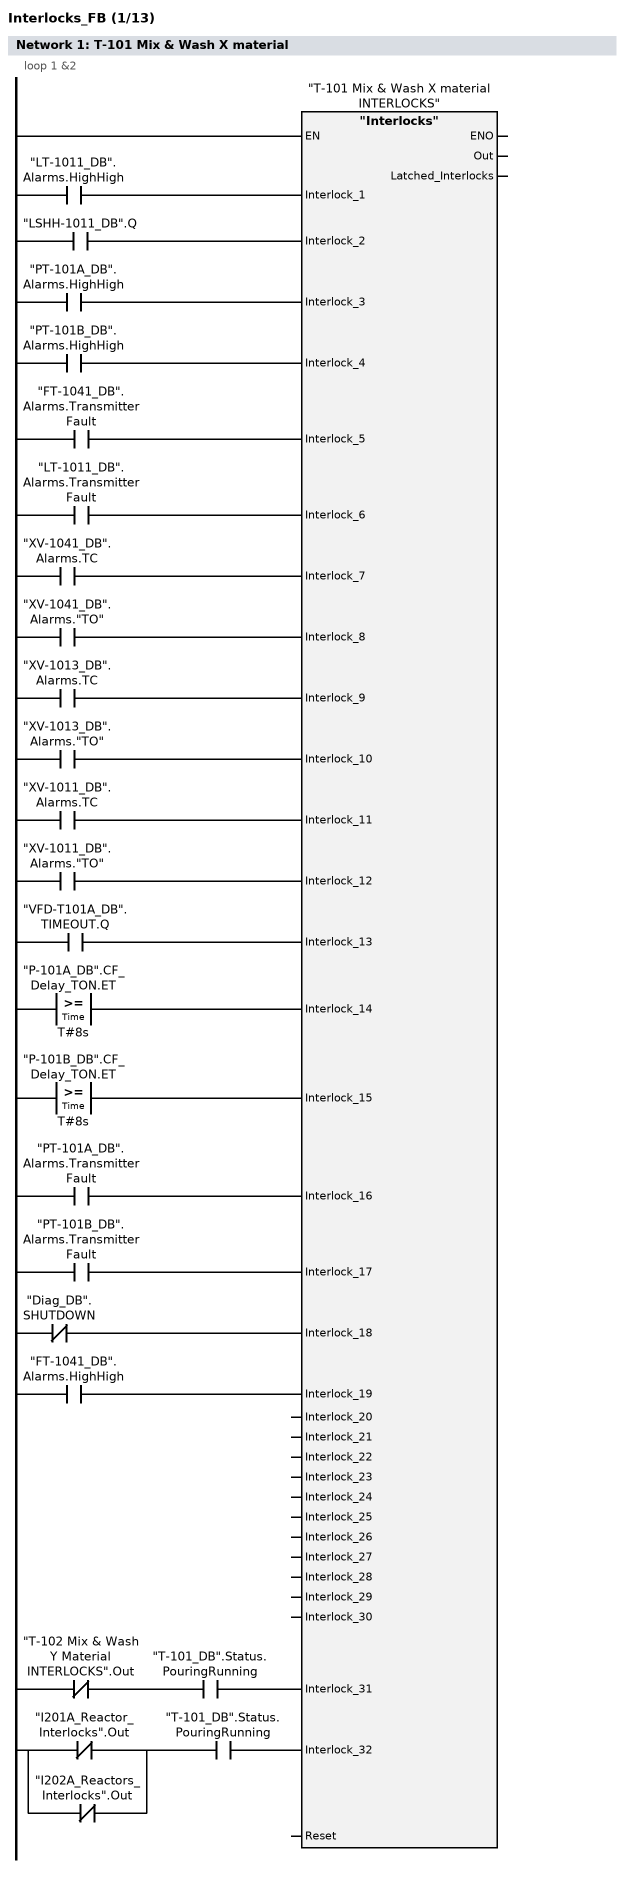
   RUNG wire#powerrail
      "T-101 Mix & Wash X material INTERLOCKS"(Interlock_1 := wire#w1, Interlock_2 := wire#w2, Interlock_3 := wire#w3, Interlock_4 := wire#w4, Interlock_5 := wire#w5, Interlock_6 := wire#w6, Interlock_7 := wire#w7, Interlock_8 := wire#w8, Interlock_9 := wire#w9, Interlock_10 := wire#w10, Interlock_11 := wire#w11, Interlock_12 := wire#w12, Interlock_13 := wire#w13, Interlock_14 := wire#w14, Interlock_15 := wire#w15, Interlock_16 := wire#w16, Interlock_17 := wire#w17, Interlock_18 := wire#w18, Interlock_19 := wire#w19, Interlock_31 := wire#w20, Interlock_32 := wire#w22, Interlock_20 :=, Interlock_21 :=, Interlock_22 :=, Interlock_23 :=, Interlock_24 :=, Interlock_25 :=, Interlock_26 :=, Interlock_27 :=, Interlock_28 :=, Interlock_29 :=, Interlock_30 :=, Reset :=, Out =>, Latched_Interlocks =>)
   END_RUNG
   RUNG wire#powerrail
      Contact( "LT-1011_DB".Alarms.HighHigh )
   END_RUNG wire#w1
   RUNG wire#powerrail
      Contact( "LSHH-1011_DB".Q )
   END_RUNG wire#w2
   RUNG wire#powerrail
      Contact( "PT-101A_DB".Alarms.HighHigh )
   END_RUNG wire#w3
   RUNG wire#powerrail
      Contact( "PT-101B_DB".Alarms.HighHigh )
   END_RUNG wire#w4
   RUNG wire#powerrail
      Contact( "FT-1041_DB".Alarms.TransmitterFault )
   END_RUNG wire#w5
   RUNG wire#powerrail
      Contact( "LT-1011_DB".Alarms.TransmitterFault )
   END_RUNG wire#w6
   RUNG wire#powerrail
      Contact( "XV-1041_DB".Alarms.TC )
   END_RUNG wire#w7
   RUNG wire#powerrail
      Contact( "XV-1041_DB".Alarms."TO" )
   END_RUNG wire#w8
   RUNG wire#powerrail
      Contact( "XV-1013_DB".Alarms.TC )
   END_RUNG wire#w9
   RUNG wire#powerrail
      Contact( "XV-1013_DB".Alarms."TO" )
   END_RUNG wire#w10
   RUNG wire#powerrail
      Contact( "XV-1011_DB".Alarms.TC )
   END_RUNG wire#w11
   RUNG wire#powerrail
      Contact( "XV-1011_DB".Alarms."TO" )
   END_RUNG wire#w12
   RUNG wire#powerrail
      Contact( "VFD-T101A_DB".TIMEOUT.Q )
   END_RUNG wire#w13
   RUNG wire#powerrail
      { S7_Templates := "SrcType := Time" } GE_Contact(in1 := "P-101A_DB".CF_Delay_TON.ET, in2 := T#8s)
   END_RUNG wire#w14
   RUNG wire#powerrail
      { S7_Templates := "SrcType := Time" } GE_Contact(in1 := "P-101B_DB".CF_Delay_TON.ET, in2 := T#8s)
   END_RUNG wire#w15
   RUNG wire#powerrail
      Contact( "PT-101A_DB".Alarms.TransmitterFault )
   END_RUNG wire#w16
   RUNG wire#powerrail
      Contact( "PT-101B_DB".Alarms.TransmitterFault )
   END_RUNG wire#w17
   RUNG wire#powerrail
      I_Contact( "Diag_DB".SHUTDOWN )
   END_RUNG wire#w18
   RUNG wire#powerrail
      Contact( "FT-1041_DB".Alarms.HighHigh )
   END_RUNG wire#w19
   RUNG wire#powerrail
      I_Contact( "T-102 Mix & Wash Y Material  INTERLOCKS".Out )
      Contact( "T-101_DB".Status.PouringRunning )
   END_RUNG wire#w20
   RUNG wire#powerrail
      I_Contact( "I201A_Reactor_Interlocks".Out )
      wire#w21
      Contact( "T-101_DB".Status.PouringRunning )
   END_RUNG wire#w22
   RUNG wire#powerrail
      I_Contact( "I202A_Reactors_Interlocks".Out )
   END_RUNG wire#w21
   // the same network as SCL:
   "T-101 Mix & Wash X material INTERLOCKS"(Interlock_1 := "LT-1011_DB".Alarms.HighHigh,   // "Interlocks"
                           Interlock_2 := "LSHH-1011_DB".Q,
                           Interlock_3 := "PT-101A_DB".Alarms.HighHigh,
                           Interlock_4 := "PT-101B_DB".Alarms.HighHigh,
                           Interlock_5 := "FT-1041_DB".Alarms.TransmitterFault,
                           Interlock_6 := "LT-1011_DB".Alarms.TransmitterFault,
                           Interlock_7 := "XV-1041_DB".Alarms.TC,
                           Interlock_8 := "XV-1041_DB".Alarms."TO",
                           Interlock_9 := "XV-1013_DB".Alarms.TC,
                           Interlock_10 := "XV-1013_DB".Alarms."TO",
                           Interlock_11 := "XV-1011_DB".Alarms.TC,
                           Interlock_12 := "XV-1011_DB".Alarms."TO",
                           Interlock_13 := "VFD-T101A_DB".TIMEOUT.Q,
                           Interlock_14 := "P-101A_DB".CF_Delay_TON.ET >= T#8s,
                           Interlock_15 := "P-101B_DB".CF_Delay_TON.ET >= T#8s,
                           Interlock_16 := "PT-101A_DB".Alarms.TransmitterFault,
                           Interlock_17 := "PT-101B_DB".Alarms.TransmitterFault,
                           Interlock_18 := NOT "Diag_DB".SHUTDOWN,
                           Interlock_19 := "FT-1041_DB".Alarms.HighHigh,
                           Interlock_31 := NOT "T-102 Mix & Wash Y Material  INTERLOCKS".Out AND "T-101_DB".Status.PouringRunning,
                           Interlock_32 := (NOT "I201A_Reactor_Interlocks".Out OR NOT "I202A_Reactors_Interlocks".Out) AND "T-101_DB".Status.PouringRunning);
END_REGION

REGION Network 2: T-102 Mix & Wash Y Material
   // loop 1 &2
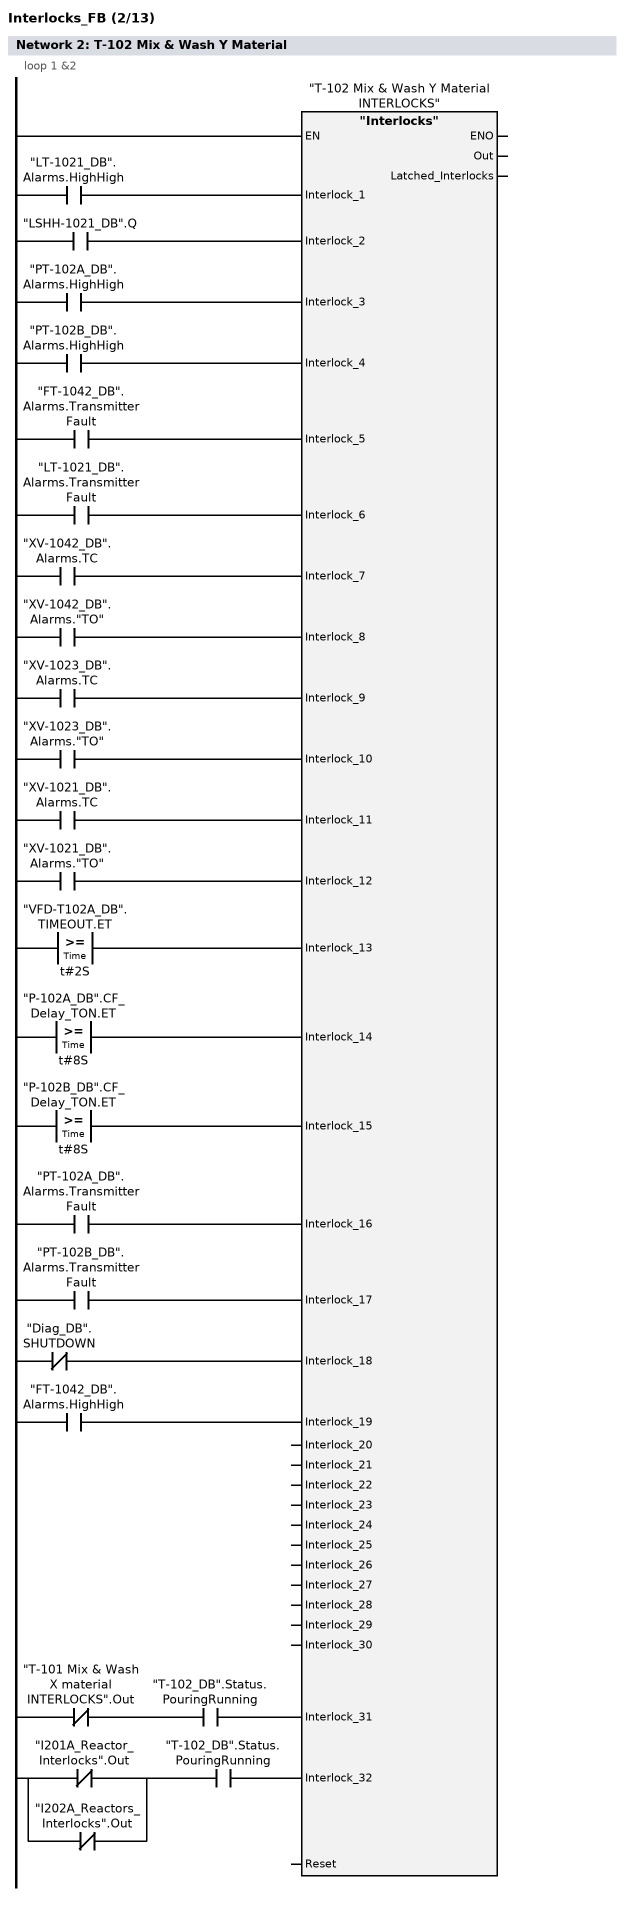
   RUNG wire#powerrail
      "T-102 Mix & Wash Y Material  INTERLOCKS"(Interlock_1 := wire#w1, Interlock_2 := wire#w2, Interlock_3 := wire#w3, Interlock_4 := wire#w4, Interlock_5 := wire#w5, Interlock_6 := wire#w6, Interlock_7 := wire#w7, Interlock_8 := wire#w8, Interlock_9 := wire#w9, Interlock_10 := wire#w10, Interlock_11 := wire#w11, Interlock_12 := wire#w12, Interlock_13 := wire#w13, Interlock_14 := wire#w14, Interlock_15 := wire#w15, Interlock_16 := wire#w16, Interlock_17 := wire#w17, Interlock_18 := wire#w18, Interlock_19 := wire#w19, Interlock_31 := wire#w20, Interlock_32 := wire#w22, Interlock_20 :=, Interlock_21 :=, Interlock_22 :=, Interlock_23 :=, Interlock_24 :=, Interlock_25 :=, Interlock_26 :=, Interlock_27 :=, Interlock_28 :=, Interlock_29 :=, Interlock_30 :=, Reset :=, Out =>, Latched_Interlocks =>)
   END_RUNG
   RUNG wire#powerrail
      Contact( "LT-1021_DB".Alarms.HighHigh )
   END_RUNG wire#w1
   RUNG wire#powerrail
      Contact( "LSHH-1021_DB".Q )
   END_RUNG wire#w2
   RUNG wire#powerrail
      Contact( "PT-102A_DB".Alarms.HighHigh )
   END_RUNG wire#w3
   RUNG wire#powerrail
      Contact( "PT-102B_DB".Alarms.HighHigh )
   END_RUNG wire#w4
   RUNG wire#powerrail
      Contact( "FT-1042_DB".Alarms.TransmitterFault )
   END_RUNG wire#w5
   RUNG wire#powerrail
      Contact( "LT-1021_DB".Alarms.TransmitterFault )
   END_RUNG wire#w6
   RUNG wire#powerrail
      Contact( "XV-1042_DB".Alarms.TC )
   END_RUNG wire#w7
   RUNG wire#powerrail
      Contact( "XV-1042_DB".Alarms."TO" )
   END_RUNG wire#w8
   RUNG wire#powerrail
      Contact( "XV-1023_DB".Alarms.TC )
   END_RUNG wire#w9
   RUNG wire#powerrail
      Contact( "XV-1023_DB".Alarms."TO" )
   END_RUNG wire#w10
   RUNG wire#powerrail
      Contact( "XV-1021_DB".Alarms.TC )
   END_RUNG wire#w11
   RUNG wire#powerrail
      Contact( "XV-1021_DB".Alarms."TO" )
   END_RUNG wire#w12
   RUNG wire#powerrail
      { S7_Templates := "SrcType := Time" } GE_Contact(in1 := "VFD-T102A_DB".TIMEOUT.ET, in2 := t#2S)
   END_RUNG wire#w13
   RUNG wire#powerrail
      { S7_Templates := "SrcType := Time" } GE_Contact(in1 := "P-102A_DB".CF_Delay_TON.ET, in2 := t#8S)
   END_RUNG wire#w14
   RUNG wire#powerrail
      { S7_Templates := "SrcType := Time" } GE_Contact(in1 := "P-102B_DB".CF_Delay_TON.ET, in2 := t#8S)
   END_RUNG wire#w15
   RUNG wire#powerrail
      Contact( "PT-102A_DB".Alarms.TransmitterFault )
   END_RUNG wire#w16
   RUNG wire#powerrail
      Contact( "PT-102B_DB".Alarms.TransmitterFault )
   END_RUNG wire#w17
   RUNG wire#powerrail
      I_Contact( "Diag_DB".SHUTDOWN )
   END_RUNG wire#w18
   RUNG wire#powerrail
      Contact( "FT-1042_DB".Alarms.HighHigh )
   END_RUNG wire#w19
   RUNG wire#powerrail
      I_Contact( "T-101 Mix & Wash X material INTERLOCKS".Out )
      Contact( "T-102_DB".Status.PouringRunning )
   END_RUNG wire#w20
   RUNG wire#powerrail
      I_Contact( "I201A_Reactor_Interlocks".Out )
      wire#w21
      Contact( "T-102_DB".Status.PouringRunning )
   END_RUNG wire#w22
   RUNG wire#powerrail
      I_Contact( "I202A_Reactors_Interlocks".Out )
   END_RUNG wire#w21
   // the same network as SCL:
   "T-102 Mix & Wash Y Material  INTERLOCKS"(Interlock_1 := "LT-1021_DB".Alarms.HighHigh,   // "Interlocks"
                           Interlock_2 := "LSHH-1021_DB".Q,
                           Interlock_3 := "PT-102A_DB".Alarms.HighHigh,
                           Interlock_4 := "PT-102B_DB".Alarms.HighHigh,
                           Interlock_5 := "FT-1042_DB".Alarms.TransmitterFault,
                           Interlock_6 := "LT-1021_DB".Alarms.TransmitterFault,
                           Interlock_7 := "XV-1042_DB".Alarms.TC,
                           Interlock_8 := "XV-1042_DB".Alarms."TO",
                           Interlock_9 := "XV-1023_DB".Alarms.TC,
                           Interlock_10 := "XV-1023_DB".Alarms."TO",
                           Interlock_11 := "XV-1021_DB".Alarms.TC,
                           Interlock_12 := "XV-1021_DB".Alarms."TO",
                           Interlock_13 := "VFD-T102A_DB".TIMEOUT.ET >= t#2S,
                           Interlock_14 := "P-102A_DB".CF_Delay_TON.ET >= t#8S,
                           Interlock_15 := "P-102B_DB".CF_Delay_TON.ET >= t#8S,
                           Interlock_16 := "PT-102A_DB".Alarms.TransmitterFault,
                           Interlock_17 := "PT-102B_DB".Alarms.TransmitterFault,
                           Interlock_18 := NOT "Diag_DB".SHUTDOWN,
                           Interlock_19 := "FT-1042_DB".Alarms.HighHigh,
                           Interlock_31 := NOT "T-101 Mix & Wash X material INTERLOCKS".Out AND "T-102_DB".Status.PouringRunning,
                           Interlock_32 := (NOT "I201A_Reactor_Interlocks".Out OR NOT "I202A_Reactors_Interlocks".Out) AND "T-102_DB".Status.PouringRunning);
END_REGION

REGION Network 3: C-301 Centrifuge interlocks
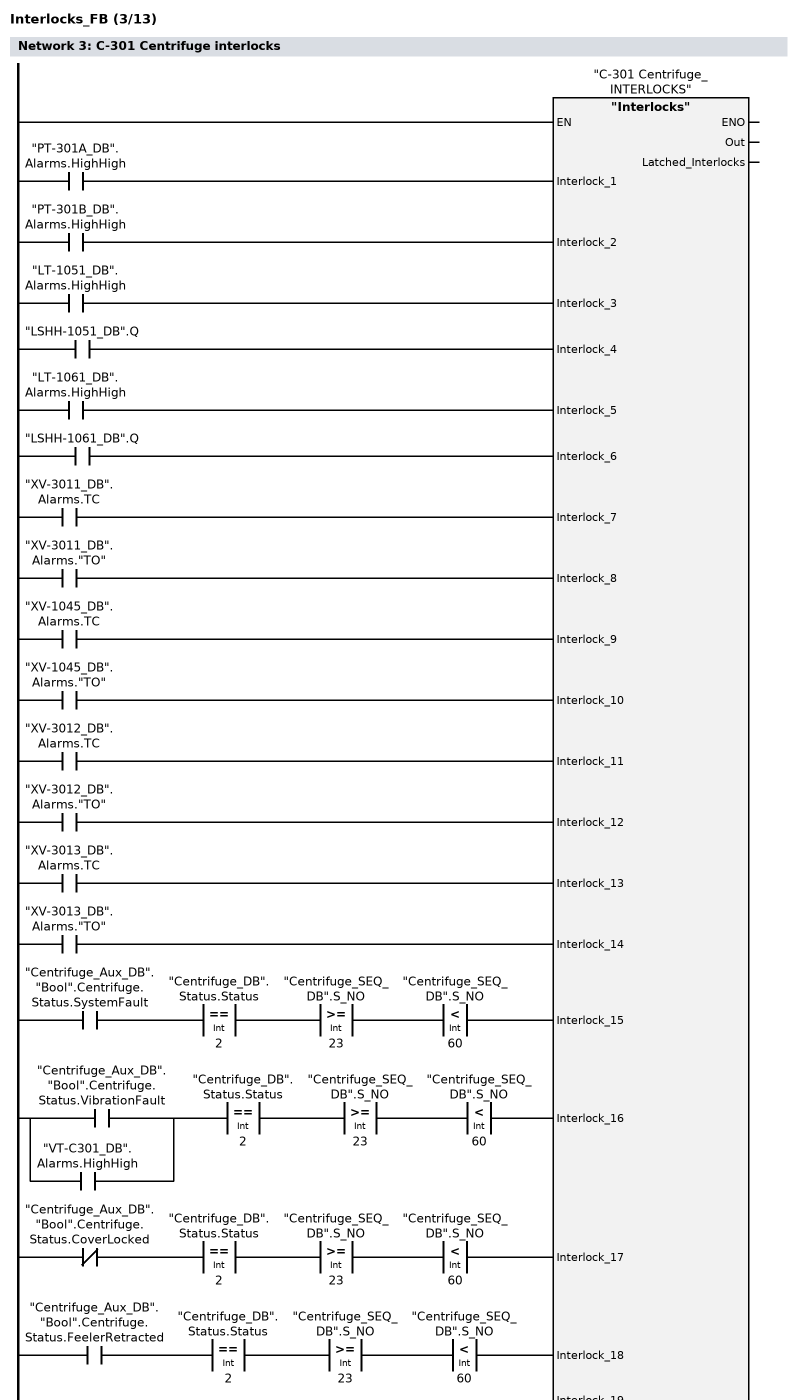
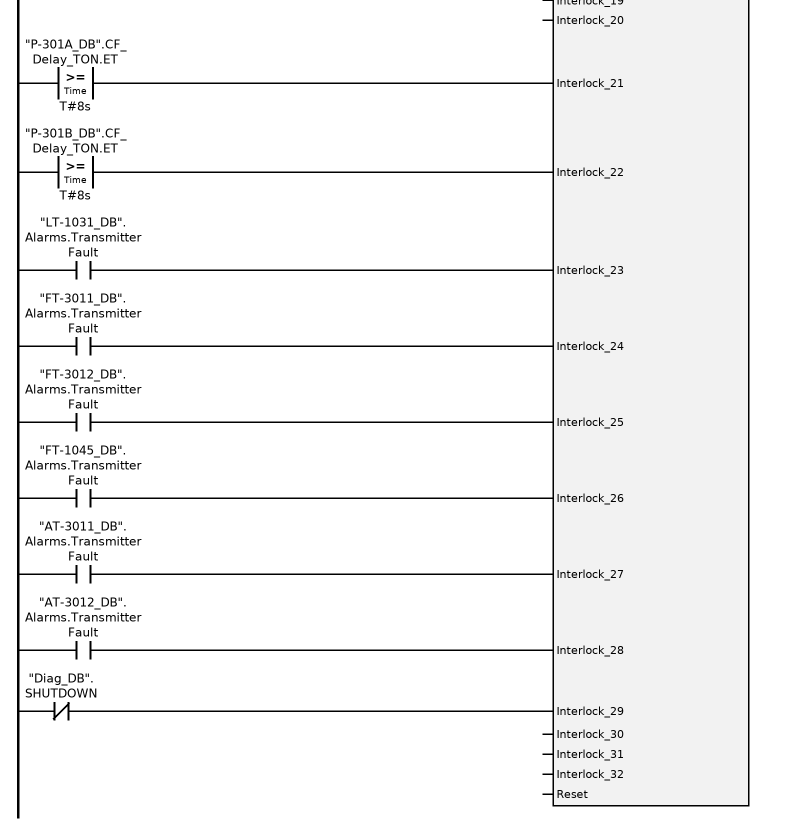
   RUNG wire#powerrail
      "C-301 Centrifuge_INTERLOCKS"(Interlock_1 := wire#w1, Interlock_2 := wire#w2, Interlock_3 := wire#w3, Interlock_4 := wire#w4, Interlock_5 := wire#w5, Interlock_6 := wire#w6, Interlock_7 := wire#w7, Interlock_8 := wire#w8, Interlock_9 := wire#w9, Interlock_10 := wire#w10, Interlock_11 := wire#w11, Interlock_12 := wire#w12, Interlock_13 := wire#w13, Interlock_14 := wire#w14, Interlock_15 := wire#w15, Interlock_16 := wire#w17, Interlock_17 := wire#w18, Interlock_18 := wire#w19, Interlock_21 := wire#w20, Interlock_22 := wire#w21, Interlock_23 := wire#w22, Interlock_24 := wire#w23, Interlock_25 := wire#w24, Interlock_26 := wire#w25, Interlock_27 := wire#w26, Interlock_28 := wire#w27, Interlock_29 := wire#w28, Interlock_19 :=, Interlock_20 :=, Interlock_30 :=, Interlock_31 :=, Interlock_32 :=, Reset :=, Out =>, Latched_Interlocks =>)
   END_RUNG
   RUNG wire#powerrail
      Contact( "PT-301A_DB".Alarms.HighHigh )
   END_RUNG wire#w1
   RUNG wire#powerrail
      Contact( "PT-301B_DB".Alarms.HighHigh )
   END_RUNG wire#w2
   RUNG wire#powerrail
      Contact( "LT-1051_DB".Alarms.HighHigh )
   END_RUNG wire#w3
   RUNG wire#powerrail
      Contact( "LSHH-1051_DB".Q )
   END_RUNG wire#w4
   RUNG wire#powerrail
      Contact( "LT-1061_DB".Alarms.HighHigh )
   END_RUNG wire#w5
   RUNG wire#powerrail
      Contact( "LSHH-1061_DB".Q )
   END_RUNG wire#w6
   RUNG wire#powerrail
      Contact( "XV-3011_DB".Alarms.TC )
   END_RUNG wire#w7
   RUNG wire#powerrail
      Contact( "XV-3011_DB".Alarms."TO" )
   END_RUNG wire#w8
   RUNG wire#powerrail
      Contact( "XV-1045_DB".Alarms.TC )
   END_RUNG wire#w9
   RUNG wire#powerrail
      Contact( "XV-1045_DB".Alarms."TO" )
   END_RUNG wire#w10
   RUNG wire#powerrail
      Contact( "XV-3012_DB".Alarms.TC )
   END_RUNG wire#w11
   RUNG wire#powerrail
      Contact( "XV-3012_DB".Alarms."TO" )
   END_RUNG wire#w12
   RUNG wire#powerrail
      Contact( "XV-3013_DB".Alarms.TC )
   END_RUNG wire#w13
   RUNG wire#powerrail
      Contact( "XV-3013_DB".Alarms."TO" )
   END_RUNG wire#w14
   RUNG wire#powerrail
      Contact( "Centrifuge_Aux_DB"."Bool".Centrifuge.Status.SystemFault )
      { S7_Templates := "SrcType := Int" } EQ_Contact(in1 := "Centrifuge_DB".Status.Status, in2 := 2)
      { S7_Templates := "SrcType := Int" } GE_Contact(in1 := "Centrifuge_SEQ_DB".S_NO, in2 := 23)
      { S7_Templates := "SrcType := Int" } LT_Contact(in1 := "Centrifuge_SEQ_DB".S_NO, in2 := 60)
   END_RUNG wire#w15
   RUNG wire#powerrail
      Contact( "Centrifuge_Aux_DB"."Bool".Centrifuge.Status.VibrationFault )
      wire#w16
      { S7_Templates := "SrcType := Int" } EQ_Contact(in1 := "Centrifuge_DB".Status.Status, in2 := 2)
      { S7_Templates := "SrcType := Int" } GE_Contact(in1 := "Centrifuge_SEQ_DB".S_NO, in2 := 23)
      { S7_Templates := "SrcType := Int" } LT_Contact(in1 := "Centrifuge_SEQ_DB".S_NO, in2 := 60)
   END_RUNG wire#w17
   RUNG wire#powerrail
      Contact( "VT-C301_DB".Alarms.HighHigh )
   END_RUNG wire#w16
   RUNG wire#powerrail
      I_Contact( "Centrifuge_Aux_DB"."Bool".Centrifuge.Status.CoverLocked )
      { S7_Templates := "SrcType := Int" } EQ_Contact(in1 := "Centrifuge_DB".Status.Status, in2 := 2)
      { S7_Templates := "SrcType := Int" } GE_Contact(in1 := "Centrifuge_SEQ_DB".S_NO, in2 := 23)
      { S7_Templates := "SrcType := Int" } LT_Contact(in1 := "Centrifuge_SEQ_DB".S_NO, in2 := 60)
   END_RUNG wire#w18
   RUNG wire#powerrail
      Contact( "Centrifuge_Aux_DB"."Bool".Centrifuge.Status.FeelerRetracted )
      { S7_Templates := "SrcType := Int" } EQ_Contact(in1 := "Centrifuge_DB".Status.Status, in2 := 2)
      { S7_Templates := "SrcType := Int" } GE_Contact(in1 := "Centrifuge_SEQ_DB".S_NO, in2 := 23)
      { S7_Templates := "SrcType := Int" } LT_Contact(in1 := "Centrifuge_SEQ_DB".S_NO, in2 := 60)
   END_RUNG wire#w19
   RUNG wire#powerrail
      { S7_Templates := "SrcType := Time" } GE_Contact(in1 := "P-301A_DB".CF_Delay_TON.ET, in2 := T#8s)
   END_RUNG wire#w20
   RUNG wire#powerrail
      { S7_Templates := "SrcType := Time" } GE_Contact(in1 := "P-301B_DB".CF_Delay_TON.ET, in2 := T#8s)
   END_RUNG wire#w21
   RUNG wire#powerrail
      Contact( "LT-1031_DB".Alarms.TransmitterFault )
   END_RUNG wire#w22
   RUNG wire#powerrail
      Contact( "FT-3011_DB".Alarms.TransmitterFault )
   END_RUNG wire#w23
   RUNG wire#powerrail
      Contact( "FT-3012_DB".Alarms.TransmitterFault )
   END_RUNG wire#w24
   RUNG wire#powerrail
      Contact( "FT-1045_DB".Alarms.TransmitterFault )
   END_RUNG wire#w25
   RUNG wire#powerrail
      Contact( "AT-3011_DB".Alarms.TransmitterFault )
   END_RUNG wire#w26
   RUNG wire#powerrail
      Contact( "AT-3012_DB".Alarms.TransmitterFault )
   END_RUNG wire#w27
   RUNG wire#powerrail
      I_Contact( "Diag_DB".SHUTDOWN )
   END_RUNG wire#w28
   // the same network as SCL:
   "C-301 Centrifuge_INTERLOCKS"(Interlock_1 := "PT-301A_DB".Alarms.HighHigh,   // "Interlocks"
                           Interlock_2 := "PT-301B_DB".Alarms.HighHigh,
                           Interlock_3 := "LT-1051_DB".Alarms.HighHigh,
                           Interlock_4 := "LSHH-1051_DB".Q,
                           Interlock_5 := "LT-1061_DB".Alarms.HighHigh,
                           Interlock_6 := "LSHH-1061_DB".Q,
                           Interlock_7 := "XV-3011_DB".Alarms.TC,
                           Interlock_8 := "XV-3011_DB".Alarms."TO",
                           Interlock_9 := "XV-1045_DB".Alarms.TC,
                           Interlock_10 := "XV-1045_DB".Alarms."TO",
                           Interlock_11 := "XV-3012_DB".Alarms.TC,
                           Interlock_12 := "XV-3012_DB".Alarms."TO",
                           Interlock_13 := "XV-3013_DB".Alarms.TC,
                           Interlock_14 := "XV-3013_DB".Alarms."TO",
                           Interlock_15 := "Centrifuge_Aux_DB"."Bool".Centrifuge.Status.SystemFault AND ("Centrifuge_DB".Status.Status = 2) AND ("Centrifuge_SEQ_DB".S_NO >= 23) AND ("Centrifuge_SEQ_DB".S_NO < 60),
                           Interlock_16 := ("Centrifuge_Aux_DB"."Bool".Centrifuge.Status.VibrationFault OR "VT-C301_DB".Alarms.HighHigh) AND ("Centrifuge_DB".Status.Status = 2) AND ("Centrifuge_SEQ_DB".S_NO >= 23) AND ("Centrifuge_SEQ_DB".S_NO < 60),
                           Interlock_17 := NOT "Centrifuge_Aux_DB"."Bool".Centrifuge.Status.CoverLocked AND ("Centrifuge_DB".Status.Status = 2) AND ("Centrifuge_SEQ_DB".S_NO >= 23) AND ("Centrifuge_SEQ_DB".S_NO < 60),
                           Interlock_18 := "Centrifuge_Aux_DB"."Bool".Centrifuge.Status.FeelerRetracted AND ("Centrifuge_DB".Status.Status = 2) AND ("Centrifuge_SEQ_DB".S_NO >= 23) AND ("Centrifuge_SEQ_DB".S_NO < 60),
                           Interlock_21 := "P-301A_DB".CF_Delay_TON.ET >= T#8s,
                           Interlock_22 := "P-301B_DB".CF_Delay_TON.ET >= T#8s,
                           Interlock_23 := "LT-1031_DB".Alarms.TransmitterFault,
                           Interlock_24 := "FT-3011_DB".Alarms.TransmitterFault,
                           Interlock_25 := "FT-3012_DB".Alarms.TransmitterFault,
                           Interlock_26 := "FT-1045_DB".Alarms.TransmitterFault,
                           Interlock_27 := "AT-3011_DB".Alarms.TransmitterFault,
                           Interlock_28 := "AT-3012_DB".Alarms.TransmitterFault,
                           Interlock_29 := NOT "Diag_DB".SHUTDOWN);
END_REGION

REGION Network 4: Calcination Interlocks (Control Loop 7)
   // Will need to add the communication fault for the EuroTherm Controller
   // Will need to add the communication fault for the Mass Flow Controller
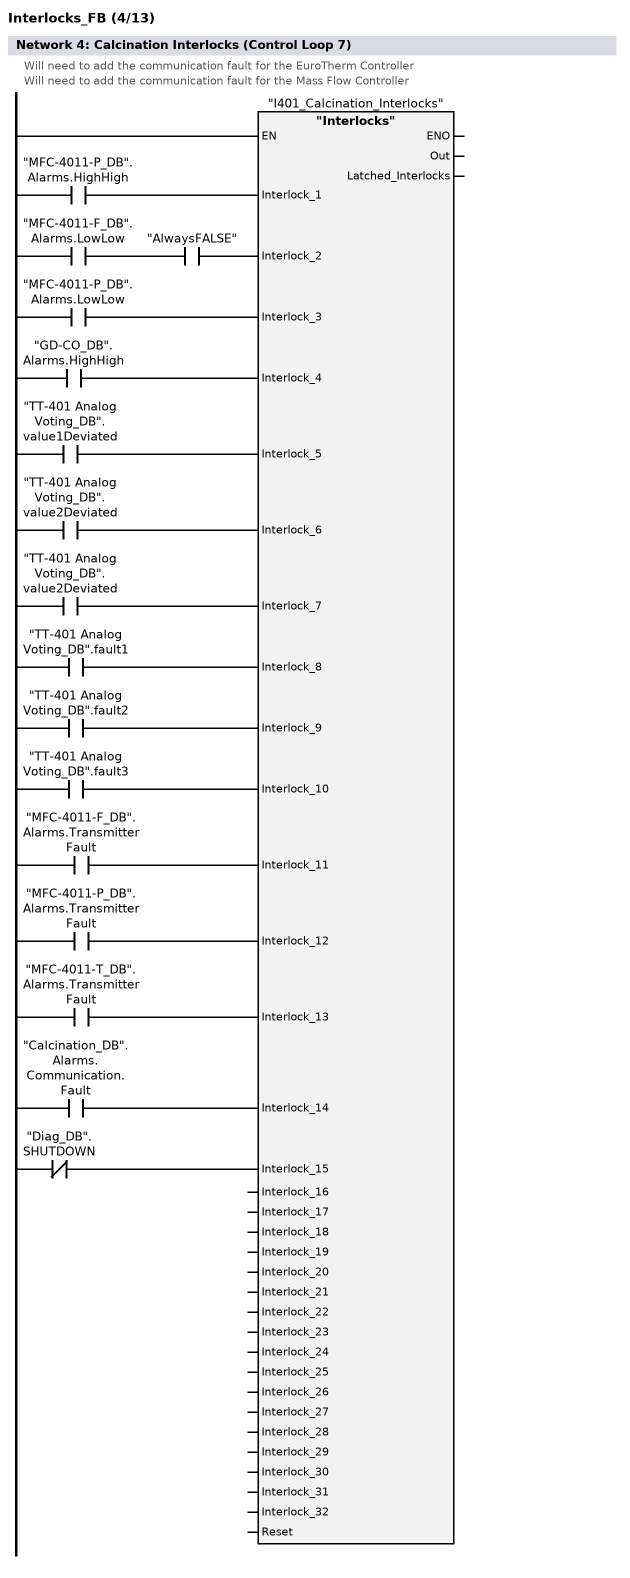
   RUNG wire#powerrail
      "I401_Calcination_Interlocks"(Interlock_1 := wire#w1, Interlock_2 := wire#w2, Interlock_3 := wire#w3, Interlock_4 := wire#w4, Interlock_5 := wire#w5, Interlock_6 := wire#w6, Interlock_7 := wire#w7, Interlock_8 := wire#w8, Interlock_9 := wire#w9, Interlock_10 := wire#w10, Interlock_11 := wire#w11, Interlock_12 := wire#w12, Interlock_13 := wire#w13, Interlock_14 := wire#w14, Interlock_15 := wire#w15, Interlock_16 :=, Interlock_17 :=, Interlock_18 :=, Interlock_19 :=, Interlock_20 :=, Interlock_21 :=, Interlock_22 :=, Interlock_23 :=, Interlock_24 :=, Interlock_25 :=, Interlock_26 :=, Interlock_27 :=, Interlock_28 :=, Interlock_29 :=, Interlock_30 :=, Interlock_31 :=, Interlock_32 :=, Reset :=, Out =>, Latched_Interlocks =>)
   END_RUNG
   RUNG wire#powerrail
      Contact( "MFC-4011-P_DB".Alarms.HighHigh )
   END_RUNG wire#w1
   RUNG wire#powerrail
      Contact( "MFC-4011-F_DB".Alarms.LowLow )
      Contact( "AlwaysFALSE" )
   END_RUNG wire#w2
   RUNG wire#powerrail
      Contact( "MFC-4011-P_DB".Alarms.LowLow )
   END_RUNG wire#w3
   RUNG wire#powerrail
      Contact( "GD-CO_DB".Alarms.HighHigh )
   END_RUNG wire#w4
   RUNG wire#powerrail
      Contact( "TT-401 Analog Voting_DB".value1Deviated )
   END_RUNG wire#w5
   RUNG wire#powerrail
      Contact( "TT-401 Analog Voting_DB".value2Deviated )
   END_RUNG wire#w6
   RUNG wire#powerrail
      Contact( "TT-401 Analog Voting_DB".value2Deviated )
   END_RUNG wire#w7
   RUNG wire#powerrail
      Contact( "TT-401 Analog Voting_DB".fault1 )
   END_RUNG wire#w8
   RUNG wire#powerrail
      Contact( "TT-401 Analog Voting_DB".fault2 )
   END_RUNG wire#w9
   RUNG wire#powerrail
      Contact( "TT-401 Analog Voting_DB".fault3 )
   END_RUNG wire#w10
   RUNG wire#powerrail
      Contact( "MFC-4011-F_DB".Alarms.TransmitterFault )
   END_RUNG wire#w11
   RUNG wire#powerrail
      Contact( "MFC-4011-P_DB".Alarms.TransmitterFault )
   END_RUNG wire#w12
   RUNG wire#powerrail
      Contact( "MFC-4011-T_DB".Alarms.TransmitterFault )
   END_RUNG wire#w13
   RUNG wire#powerrail
      Contact( "Calcination_DB".Alarms.Communication.Fault )
   END_RUNG wire#w14
   RUNG wire#powerrail
      I_Contact( "Diag_DB".SHUTDOWN )
   END_RUNG wire#w15
   // the same network as SCL:
   "I401_Calcination_Interlocks"(Interlock_1 := "MFC-4011-P_DB".Alarms.HighHigh,   // "Interlocks"
                           Interlock_2 := "MFC-4011-F_DB".Alarms.LowLow AND "AlwaysFALSE",
                           Interlock_3 := "MFC-4011-P_DB".Alarms.LowLow,
                           Interlock_4 := "GD-CO_DB".Alarms.HighHigh,
                           Interlock_5 := "TT-401 Analog Voting_DB".value1Deviated,
                           Interlock_6 := "TT-401 Analog Voting_DB".value2Deviated,
                           Interlock_7 := "TT-401 Analog Voting_DB".value2Deviated,
                           Interlock_8 := "TT-401 Analog Voting_DB".fault1,
                           Interlock_9 := "TT-401 Analog Voting_DB".fault2,
                           Interlock_10 := "TT-401 Analog Voting_DB".fault3,
                           Interlock_11 := "MFC-4011-F_DB".Alarms.TransmitterFault,
                           Interlock_12 := "MFC-4011-P_DB".Alarms.TransmitterFault,
                           Interlock_13 := "MFC-4011-T_DB".Alarms.TransmitterFault,
                           Interlock_14 := "Calcination_DB".Alarms.Communication.Fault,
                           Interlock_15 := NOT "Diag_DB".SHUTDOWN);
END_REGION

REGION Network 5: I402 Passivate Interlocks (Control Loop 8)
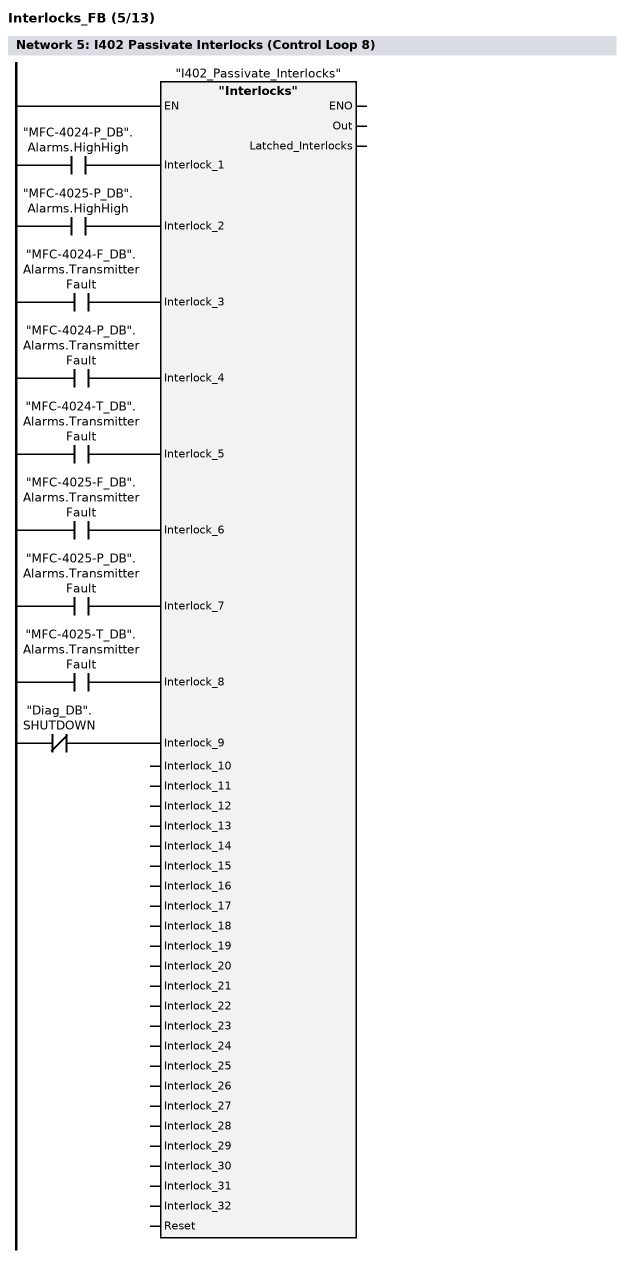
   RUNG wire#powerrail
      "I402_Passivate_Interlocks"(Interlock_1 := wire#w1, Interlock_2 := wire#w2, Interlock_3 := wire#w3, Interlock_4 := wire#w4, Interlock_5 := wire#w5, Interlock_6 := wire#w6, Interlock_7 := wire#w7, Interlock_8 := wire#w8, Interlock_9 := wire#w9, Interlock_10 :=, Interlock_11 :=, Interlock_12 :=, Interlock_13 :=, Interlock_14 :=, Interlock_15 :=, Interlock_16 :=, Interlock_17 :=, Interlock_18 :=, Interlock_19 :=, Interlock_20 :=, Interlock_21 :=, Interlock_22 :=, Interlock_23 :=, Interlock_24 :=, Interlock_25 :=, Interlock_26 :=, Interlock_27 :=, Interlock_28 :=, Interlock_29 :=, Interlock_30 :=, Interlock_31 :=, Interlock_32 :=, Reset :=, Out =>, Latched_Interlocks =>)
   END_RUNG
   RUNG wire#powerrail
      Contact( "MFC-4024-P_DB".Alarms.HighHigh )
   END_RUNG wire#w1
   RUNG wire#powerrail
      Contact( "MFC-4025-P_DB".Alarms.HighHigh )
   END_RUNG wire#w2
   RUNG wire#powerrail
      Contact( "MFC-4024-F_DB".Alarms.TransmitterFault )
   END_RUNG wire#w3
   RUNG wire#powerrail
      Contact( "MFC-4024-P_DB".Alarms.TransmitterFault )
   END_RUNG wire#w4
   RUNG wire#powerrail
      Contact( "MFC-4024-T_DB".Alarms.TransmitterFault )
   END_RUNG wire#w5
   RUNG wire#powerrail
      Contact( "MFC-4025-F_DB".Alarms.TransmitterFault )
   END_RUNG wire#w6
   RUNG wire#powerrail
      Contact( "MFC-4025-P_DB".Alarms.TransmitterFault )
   END_RUNG wire#w7
   RUNG wire#powerrail
      Contact( "MFC-4025-T_DB".Alarms.TransmitterFault )
   END_RUNG wire#w8
   RUNG wire#powerrail
      I_Contact( "Diag_DB".SHUTDOWN )
   END_RUNG wire#w9
   // the same network as SCL:
   "I402_Passivate_Interlocks"(Interlock_1 := "MFC-4024-P_DB".Alarms.HighHigh,   // "Interlocks"
                           Interlock_2 := "MFC-4025-P_DB".Alarms.HighHigh,
                           Interlock_3 := "MFC-4024-F_DB".Alarms.TransmitterFault,
                           Interlock_4 := "MFC-4024-P_DB".Alarms.TransmitterFault,
                           Interlock_5 := "MFC-4024-T_DB".Alarms.TransmitterFault,
                           Interlock_6 := "MFC-4025-F_DB".Alarms.TransmitterFault,
                           Interlock_7 := "MFC-4025-P_DB".Alarms.TransmitterFault,
                           Interlock_8 := "MFC-4025-T_DB".Alarms.TransmitterFault,
                           Interlock_9 := NOT "Diag_DB".SHUTDOWN);
END_REGION

REGION Network 6: I201A Reactors Interlocks (R-201)
